(* Logix 5000 project; controller PLC_MCC1201_220AP1 vendor 1 type 14 code 164 rev 35.11; software revision 35.00; part 13 of 25 *)
(* tags used below, declared in another part *)
   B180 : DINT[10];
   B3 : DINT[102];
   BIN_1B_EAST : ALIAS FOR O[112].12;
   BT181_000 : MESSAGE;
   BT181_001 : MESSAGE;
   BT181_002 : MESSAGE;
   BT181_003 : MESSAGE;
   C1_PNL_FLT : ALIAS FOR I[113].2;
   C2_PNL_FLT : ALIAS FOR I[113].3;
   C3_PNL_FLT : ALIAS FOR I[113].4;
   C4_PNL_FLT : ALIAS FOR I[113].1;
   C5 : COUNTER[100];
   CAP_ALM_HORN : ALIAS FOR O[11].2;
   CR1_DOWN_PROX : ALIAS FOR I[64].11;
   CR1_RUN_ENABLE : ALIAS FOR O[117].4;
   CULL_FLT : ALIAS FOR B3[3].1;
   CULLET_FLT_PL : ALIAS FOR O[11].1;
   DIV_POSITION : ALIAS FOR I[24].12;
   I : INT[128];
   LEG2_SLEEP : ALIAS FOR I[123].14;
   LEG3_SLEEP : ALIAS FOR I[123].15;
   LEG4_SLEEP : ALIAS FOR I[124].0;
   LEG5_SLEEP : ALIAS FOR I[124].1;
   M37B_FWD_DIR : ALIAS FOR B3[1].14;
   M37B_FWD_PL : ALIAS FOR O[25].5;
   M37B_FWD_SIG : ALIAS FOR I[112].3;
   M37B_FWD_SS : ALIAS FOR I[24].8;
   M37B_REV_DIR : ALIAS FOR B3[1].15;
   M37B_REV_PL : ALIAS FOR O[25].6;
   M37B_REV_SIG : ALIAS FOR I[112].4;
   M37B_REV_SS : ALIAS FOR I[24].9;
   M37B_RUN_FWD : ALIAS FOR O[119].0;
   M37B_RUN_REV : ALIAS FOR O[119].1;
   M47_REV_SS : ALIAS FOR I[24].11;
   M47B_FWD_DIR : ALIAS FOR B3[1].12;
   M47B_FWD_PL : ALIAS FOR O[25].7;
   M47B_FWD_SIG : ALIAS FOR I[112].1;
   M47B_FWD_SS : ALIAS FOR I[24].10;
   M47B_REV_DIR : ALIAS FOR B3[1].13;
   M47B_REV_PL : ALIAS FOR O[25].8;
   M47B_REV_SIG : ALIAS FOR I[112].2;
   M47B_RUN_FWD : ALIAS FOR O[119].2;
   M47B_RUN_REV : ALIAS FOR O[119].3;
   N53 : DINT[10];
   N54 : DINT[501];
   N60 : DINT[420];
   O : INT[128];
   REL_DRV_FLT : ALIAS FOR B3[3].0;
   RELIANCE_FLT_PL : ALIAS FOR O[11].0;
   S : INT[128];
   SPNGE_DN_FLT : ALIAS FOR I[43].5;
   SPNGE_UP_FLT : ALIAS FOR I[43].4;
   Status : INT;   // INT tag to retrieve Status value through GSV created during conversion
   T4 : TIMER[100];
   T51 : TIMER[13];
   TMP_xAlwaysOFF : BOOL;
   TONY : ALIAS FOR B3[10].15;
   VMCCMB_ALM_HRN : ALIAS FOR O[20].3;
   VP917060_MED : ALIAS FOR O[116].14;
   VP917060_THICK : ALIAS FOR O[116].15;
   VP917060_THIN : ALIAS FOR O[116].13;
   VP917065_MED : ALIAS FOR O[114].5;
   VP917065_THICK : ALIAS FOR O[114].6;
   VP917065_THIN : ALIAS FOR O[114].4;
   VP917066_MED : ALIAS FOR O[114].2;
   VP917066_THICK : ALIAS FOR O[114].3;
   VP917066_THIN : ALIAS FOR O[114].1;
   VP917067_MED : ALIAS FOR O[113].15;
   VP917067_THICK : ALIAS FOR O[114].0;
   VP917067_THIN : ALIAS FOR O[113].14;
   VP917070_MED : ALIAS FOR O[114].8;
   VP917070_THICK : ALIAS FOR O[114].9;
   VP917070_THIN : ALIAS FOR O[114].7;
   VP917071_MED : ALIAS FOR O[114].11;
   VP917071_THICK : ALIAS FOR O[114].12;
   VP917071_THIN : ALIAS FOR O[114].10;
   VP917072_MED : ALIAS FOR O[116].11;
   VP917072_THICK : ALIAS FOR O[116].12;
   VP917072_THIN : ALIAS FOR O[116].10;
   VP917073_MED : ALIAS FOR O[115].14;
   VP917073_THICK : ALIAS FOR O[115].15;
   VP917073_THIN : ALIAS FOR O[115].13;
   VP917074_MED : ALIAS FOR O[115].11;
   VP917074_THICK : ALIAS FOR O[115].12;
   VP917074_THIN : ALIAS FOR O[115].10;
   VP917075_MED : ALIAS FOR O[115].8;
   VP917075_THICK : ALIAS FOR O[115].9;
   VP917075_THIN : ALIAS FOR O[115].7;
   VP917076_MED : ALIAS FOR O[115].5;
   VP917076_THICK : ALIAS FOR O[115].6;
   VP917076_THIN : ALIAS FOR O[115].4;
   VP917077_MED : ALIAS FOR O[114].14;
   VP917077_THICK : ALIAS FOR O[114].15;
   VP917077_THIN : ALIAS FOR O[114].13;
   W1_DRV_FLT_RES : ALIAS FOR O[47].2;
(* MainProgram, continued *)

ROUTINE _107_LADDER   (* ladder *)
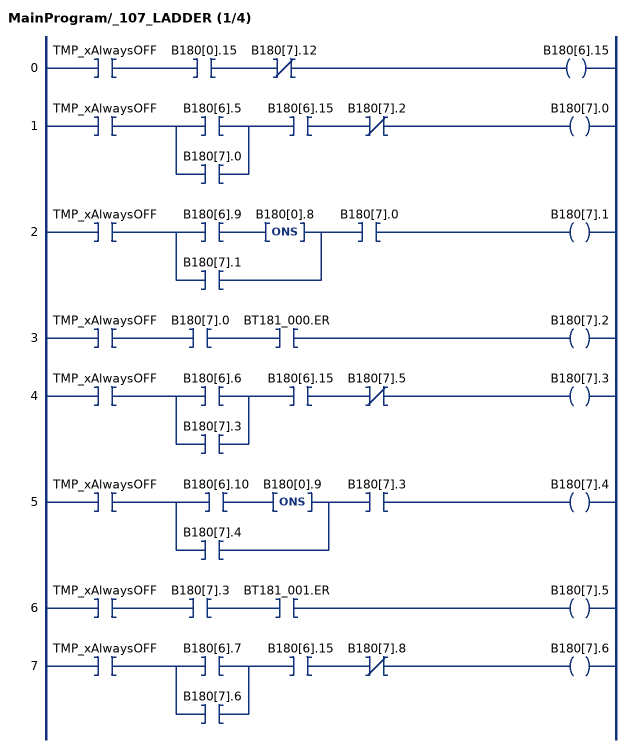
   0: XIC(TMP_xAlwaysOFF)XIC(B180[0].15)XIO(B180[7].12)OTE(B180[6].15);
   1: XIC(TMP_xAlwaysOFF)[XIC(B180[6].5) ,XIC(B180[7].0) ]XIC(B180[6].15)XIO(B180[7].2)OTE(B180[7].0);
   2: XIC(TMP_xAlwaysOFF)[XIC(B180[6].9) ONS(B180[0].8) ,XIC(B180[7].1) ]XIC(B180[7].0)OTE(B180[7].1);
   3: XIC(TMP_xAlwaysOFF)XIC(B180[7].0)XIC(BT181_000.ER)OTE(B180[7].2);
   4: XIC(TMP_xAlwaysOFF)[XIC(B180[6].6) ,XIC(B180[7].3) ]XIC(B180[6].15)XIO(B180[7].5)OTE(B180[7].3);
   5: XIC(TMP_xAlwaysOFF)[XIC(B180[6].10) ONS(B180[0].9) ,XIC(B180[7].4) ]XIC(B180[7].3)OTE(B180[7].4);
   6: XIC(TMP_xAlwaysOFF)XIC(B180[7].3)XIC(BT181_001.ER)OTE(B180[7].5);
   7: XIC(TMP_xAlwaysOFF)[XIC(B180[6].7) ,XIC(B180[7].6) ]XIC(B180[6].15)XIO(B180[7].8)OTE(B180[7].6);
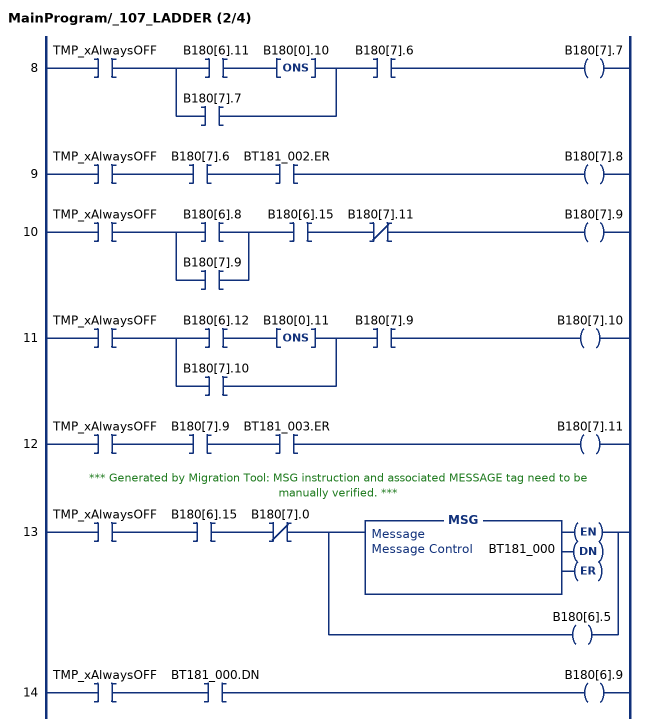
   8: XIC(TMP_xAlwaysOFF)[XIC(B180[6].11) ONS(B180[0].10) ,XIC(B180[7].7) ]XIC(B180[7].6)OTE(B180[7].7);
   9: XIC(TMP_xAlwaysOFF)XIC(B180[7].6)XIC(BT181_002.ER)OTE(B180[7].8);
   10: XIC(TMP_xAlwaysOFF)[XIC(B180[6].8) ,XIC(B180[7].9) ]XIC(B180[6].15)XIO(B180[7].11)OTE(B180[7].9);
   11: XIC(TMP_xAlwaysOFF)[XIC(B180[6].12) ONS(B180[0].11) ,XIC(B180[7].10) ]XIC(B180[7].9)OTE(B180[7].10);
   12: XIC(TMP_xAlwaysOFF)XIC(B180[7].9)XIC(BT181_003.ER)OTE(B180[7].11);
   // *** Generated by Migration Tool: MSG instruction and associated MESSAGE tag need to be manually verified. ***
   13: XIC(TMP_xAlwaysOFF)XIC(B180[6].15)XIO(B180[7].0)[MSG(BT181_000) ,OTE(B180[6].5) ];
   14: XIC(TMP_xAlwaysOFF)XIC(BT181_000.DN)OTE(B180[6].9);
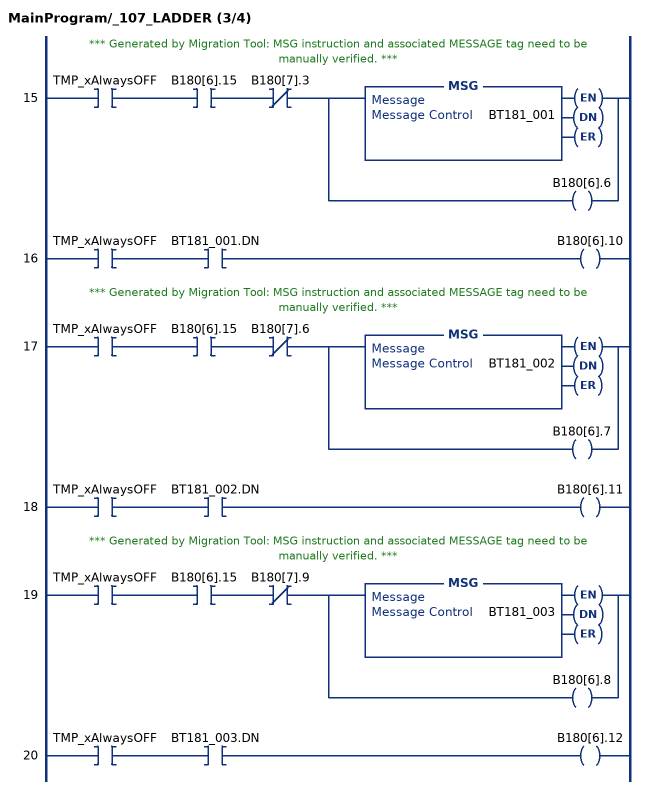
   // *** Generated by Migration Tool: MSG instruction and associated MESSAGE tag need to be manually verified. ***
   15: XIC(TMP_xAlwaysOFF)XIC(B180[6].15)XIO(B180[7].3)[MSG(BT181_001) ,OTE(B180[6].6) ];
   16: XIC(TMP_xAlwaysOFF)XIC(BT181_001.DN)OTE(B180[6].10);
   // *** Generated by Migration Tool: MSG instruction and associated MESSAGE tag need to be manually verified. ***
   17: XIC(TMP_xAlwaysOFF)XIC(B180[6].15)XIO(B180[7].6)[MSG(BT181_002) ,OTE(B180[6].7) ];
   18: XIC(TMP_xAlwaysOFF)XIC(BT181_002.DN)OTE(B180[6].11);
   // *** Generated by Migration Tool: MSG instruction and associated MESSAGE tag need to be manually verified. ***
   19: XIC(TMP_xAlwaysOFF)XIC(B180[6].15)XIO(B180[7].9)[MSG(BT181_003) ,OTE(B180[6].8) ];
   20: XIC(TMP_xAlwaysOFF)XIC(BT181_003.DN)OTE(B180[6].12);
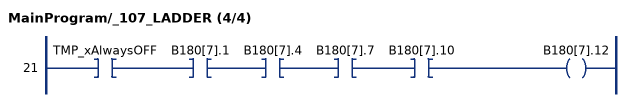
   21: XIC(TMP_xAlwaysOFF)XIC(B180[7].1)XIC(B180[7].4)XIC(B180[7].7)XIC(B180[7].10)OTE(B180[7].12);
END_ROUTINE

ROUTINE _10_SLEEP   (* ladder *)
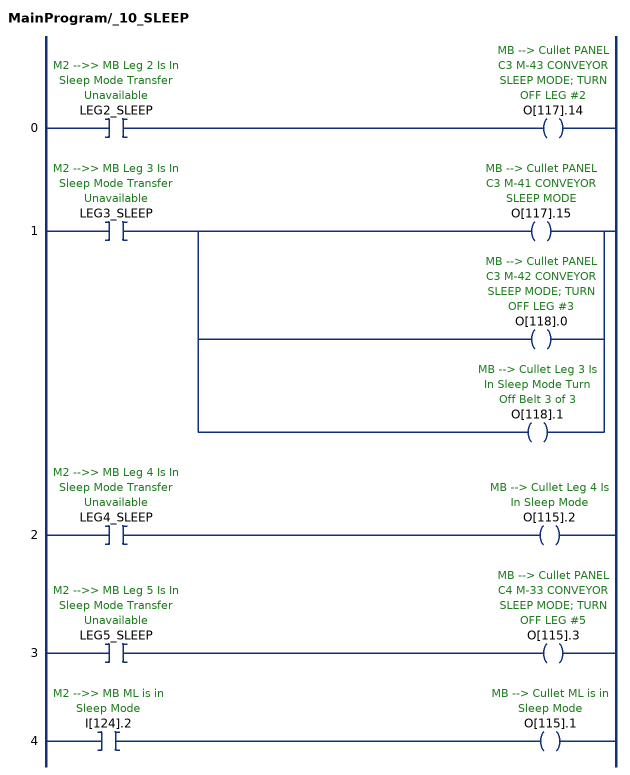
   0: XIC(LEG2_SLEEP)OTE(O[117].14);
   1: XIC(LEG3_SLEEP)[OTE(O[117].15) ,OTE(O[118].0) ,OTE(O[118].1) ];
   2: XIC(LEG4_SLEEP)OTE(O[115].2);
   3: XIC(LEG5_SLEEP)OTE(O[115].3);
   4: XIC(I[124].2)OTE(O[115].1);
END_ROUTINE

ROUTINE _11_CULLET   (* ladder *)
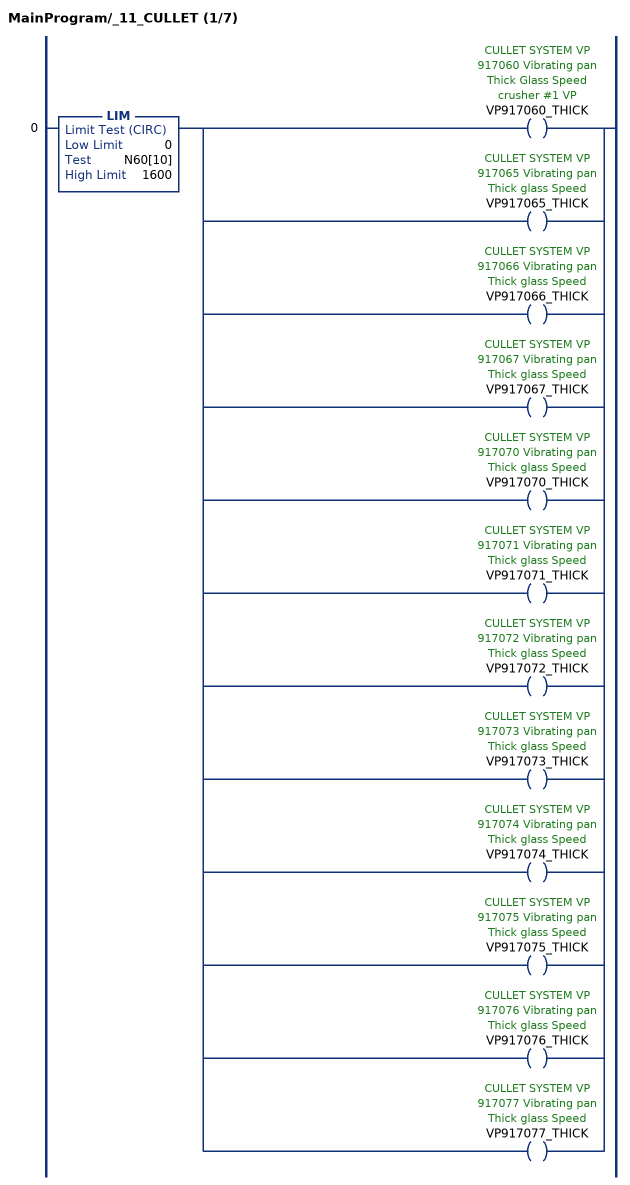
   0: LIM(0,N60[10],1600)[OTE(VP917060_THICK) ,OTE(VP917065_THICK) ,OTE(VP917066_THICK) ,OTE(VP917067_THICK) ,OTE(VP917070_THICK) ,OTE(VP917071_THICK) ,OTE(VP917072_THICK) ,OTE(VP917073_THICK) ,OTE(VP917074_THICK) ,OTE(VP917075_THICK) ,OTE(VP917076_THICK) ,OTE(VP917077_THICK) ];
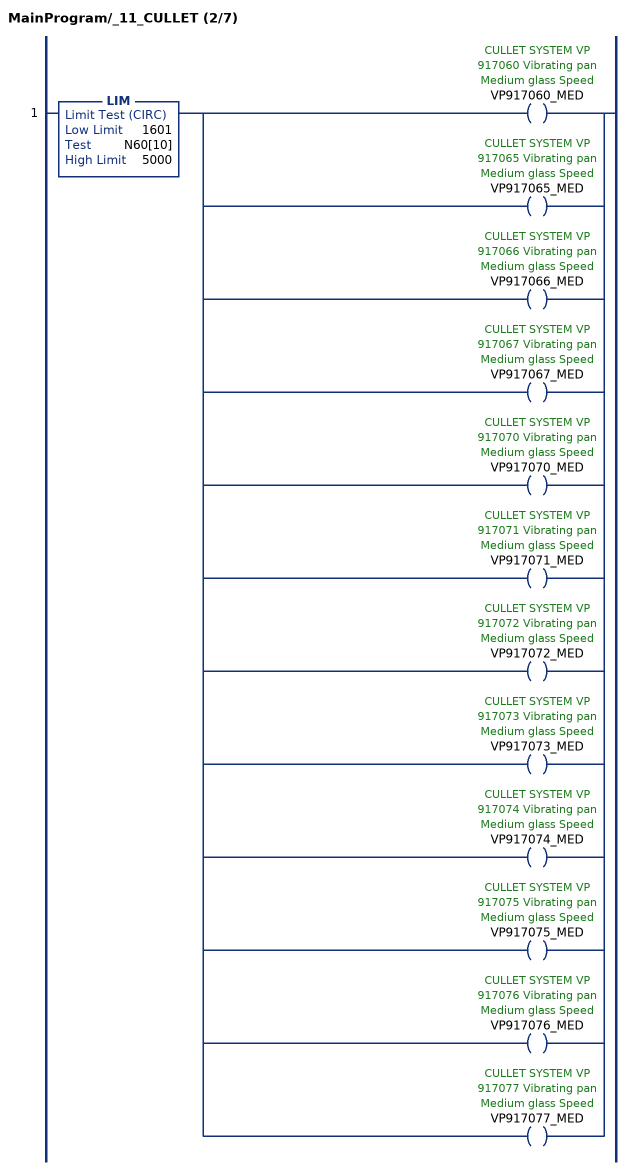
   1: LIM(1601,N60[10],5000)[OTE(VP917060_MED) ,OTE(VP917065_MED) ,OTE(VP917066_MED) ,OTE(VP917067_MED) ,OTE(VP917070_MED) ,OTE(VP917071_MED) ,OTE(VP917072_MED) ,OTE(VP917073_MED) ,OTE(VP917074_MED) ,OTE(VP917075_MED) ,OTE(VP917076_MED) ,OTE(VP917077_MED) ];
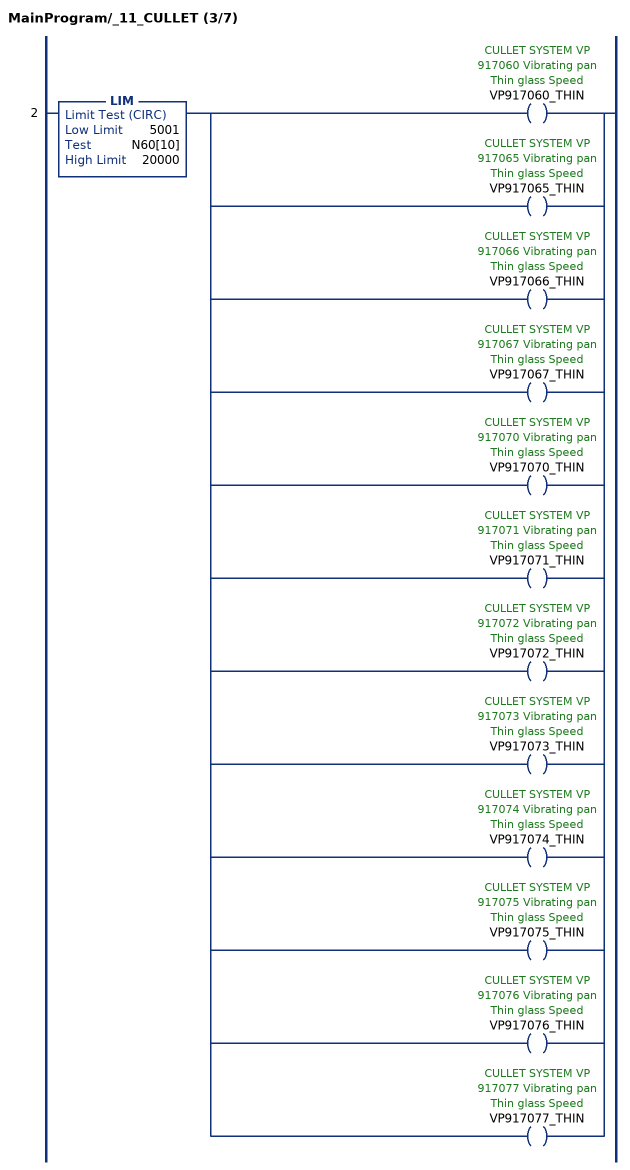
   2: LIM(5001,N60[10],20000)[OTE(VP917060_THIN) ,OTE(VP917065_THIN) ,OTE(VP917066_THIN) ,OTE(VP917067_THIN) ,OTE(VP917070_THIN) ,OTE(VP917071_THIN) ,OTE(VP917072_THIN) ,OTE(VP917073_THIN) ,OTE(VP917074_THIN) ,OTE(VP917075_THIN) ,OTE(VP917076_THIN) ,OTE(VP917077_THIN) ];
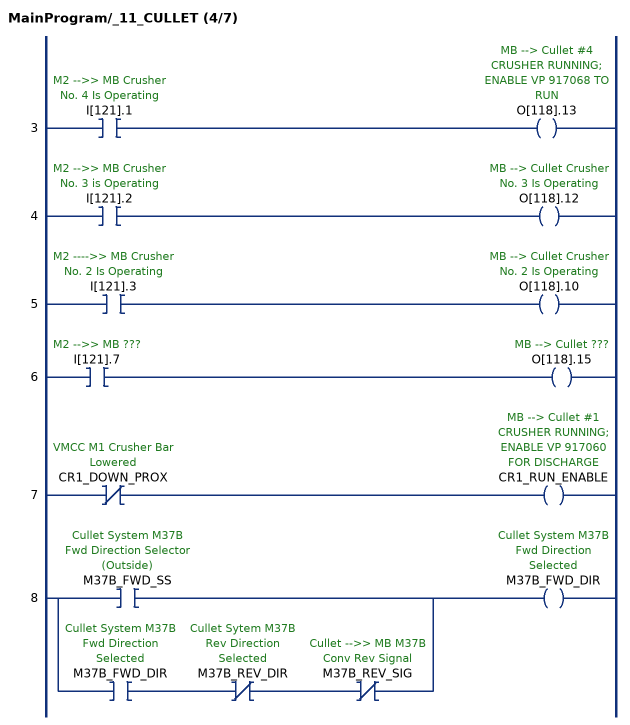
   3: XIC(I[121].1)OTE(O[118].13);
   4: XIC(I[121].2)OTE(O[118].12);
   5: XIC(I[121].3)OTE(O[118].10);
   6: XIC(I[121].7)OTE(O[118].15);
   7: XIO(CR1_DOWN_PROX)OTE(CR1_RUN_ENABLE);
   8: [XIC(M37B_FWD_SS) ,XIC(M37B_FWD_DIR) XIO(M37B_REV_DIR) XIO(M37B_REV_SIG) ]OTE(M37B_FWD_DIR);
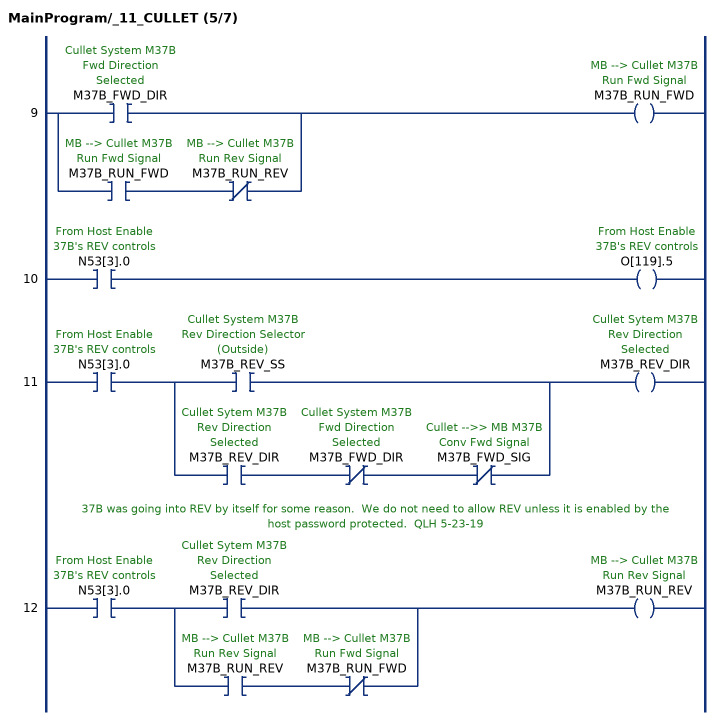
   9: [XIC(M37B_FWD_DIR) ,XIC(M37B_RUN_FWD) XIO(M37B_RUN_REV) ]OTE(M37B_RUN_FWD);
   10: XIC(N53[3].0)OTE(O[119].5);
   11: XIC(N53[3].0)[XIC(M37B_REV_SS) ,XIC(M37B_REV_DIR) XIO(M37B_FWD_DIR) XIO(M37B_FWD_SIG) ]OTE(M37B_REV_DIR);
   // 37B was going into REV by itself for some reason.  We do not need to allow REV unless it is enabled by the host password protected.  QLH 5-23-19
   12: XIC(N53[3].0)[XIC(M37B_REV_DIR) ,XIC(M37B_RUN_REV) XIO(M37B_RUN_FWD) ]OTE(M37B_RUN_REV);
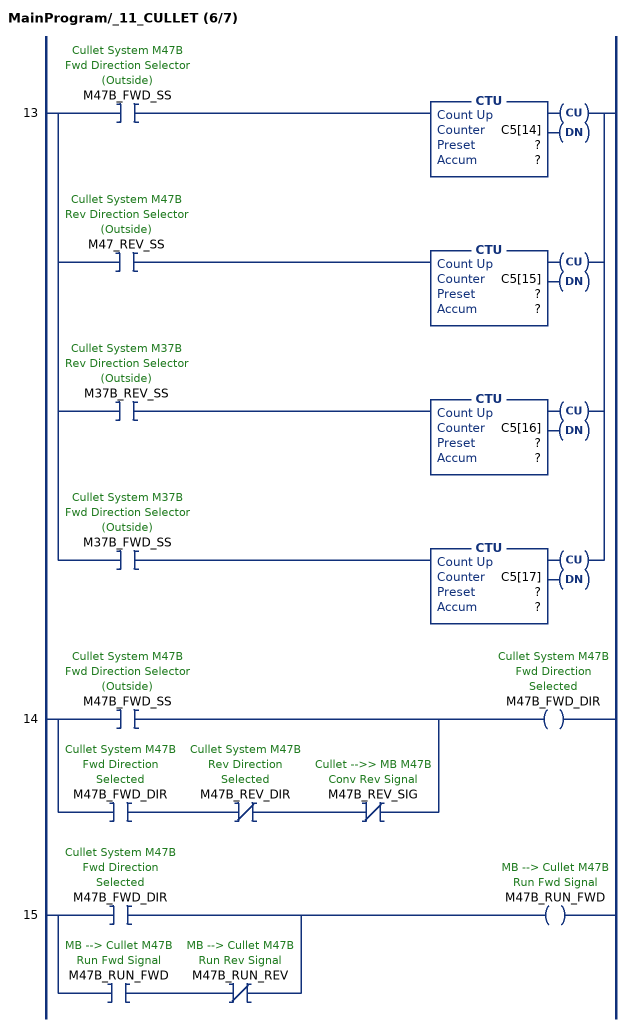
   13: [XIC(M47B_FWD_SS) CTU(C5[14],?,?) ,XIC(M47_REV_SS) CTU(C5[15],?,?) ,XIC(M37B_REV_SS) CTU(C5[16],?,?) ,XIC(M37B_FWD_SS) CTU(C5[17],?,?) ];
   14: [XIC(M47B_FWD_SS) ,XIC(M47B_FWD_DIR) XIO(M47B_REV_DIR) XIO(M47B_REV_SIG) ]OTE(M47B_FWD_DIR);
   15: [XIC(M47B_FWD_DIR) ,XIC(M47B_RUN_FWD) XIO(M47B_RUN_REV) ]OTE(M47B_RUN_FWD);
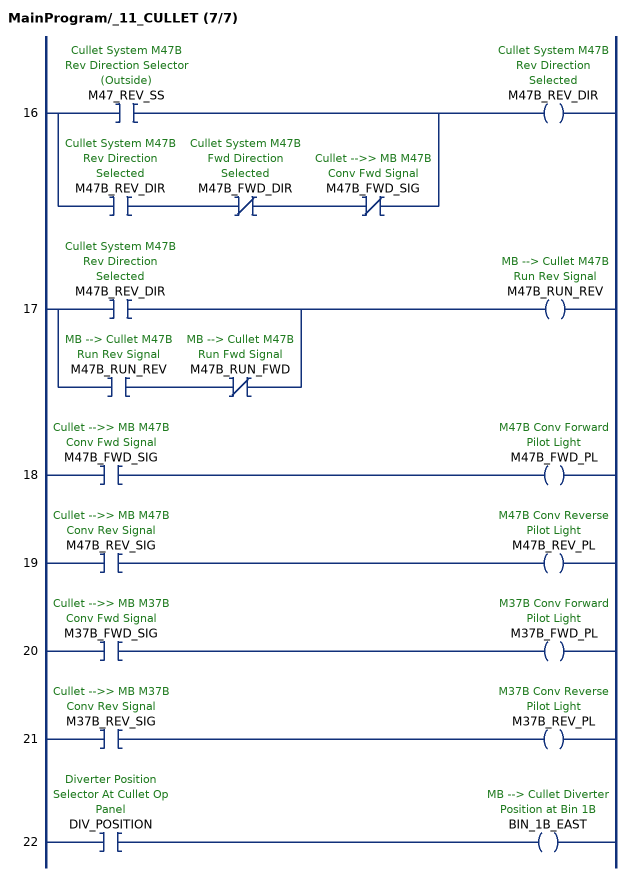
   16: [XIC(M47_REV_SS) ,XIC(M47B_REV_DIR) XIO(M47B_FWD_DIR) XIO(M47B_FWD_SIG) ]OTE(M47B_REV_DIR);
   17: [XIC(M47B_REV_DIR) ,XIC(M47B_RUN_REV) XIO(M47B_RUN_FWD) ]OTE(M47B_RUN_REV);
   18: XIC(M47B_FWD_SIG)OTE(M47B_FWD_PL);
   19: XIC(M47B_REV_SIG)OTE(M47B_REV_PL);
   20: XIC(M37B_FWD_SIG)OTE(M37B_FWD_PL);
   21: XIC(M37B_REV_SIG)OTE(M37B_REV_PL);
   22: XIC(DIV_POSITION)OTE(BIN_1B_EAST);
END_ROUTINE

ROUTINE _12_MAIN   (* ladder *)
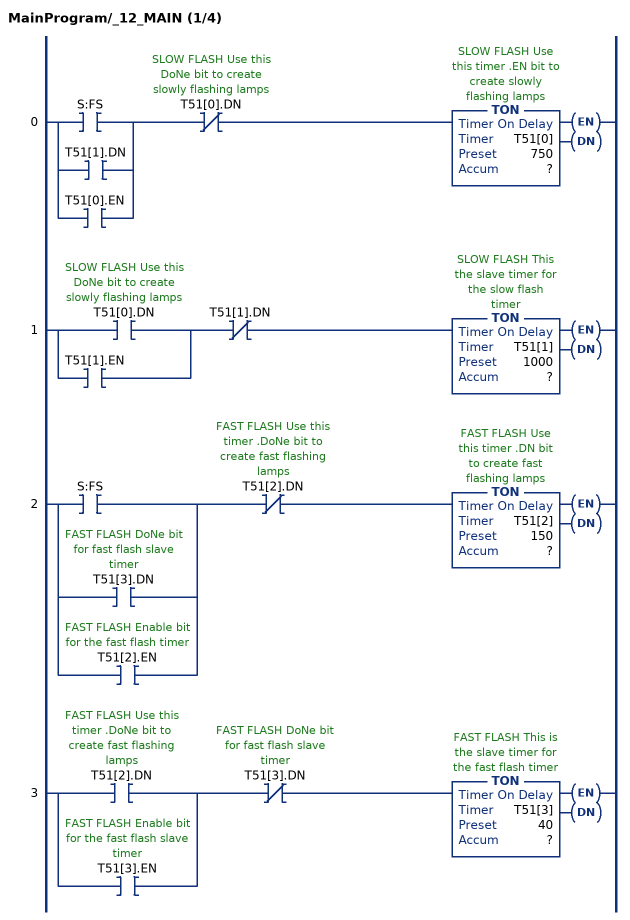
   0: [XIC(S:FS) ,XIC(T51[1].DN) ,XIC(T51[0].EN) ]XIO(T51[0].DN)TON(T51[0],?,?);
   1: [XIC(T51[0].DN) ,XIC(T51[1].EN) ]XIO(T51[1].DN)TON(T51[1],?,?);
   2: [XIC(S:FS) ,XIC(T51[3].DN) ,XIC(T51[2].EN) ]XIO(T51[2].DN)TON(T51[2],?,?);
   3: [XIC(T51[2].DN) ,XIC(T51[3].EN) ]XIO(T51[3].DN)TON(T51[3],?,?);
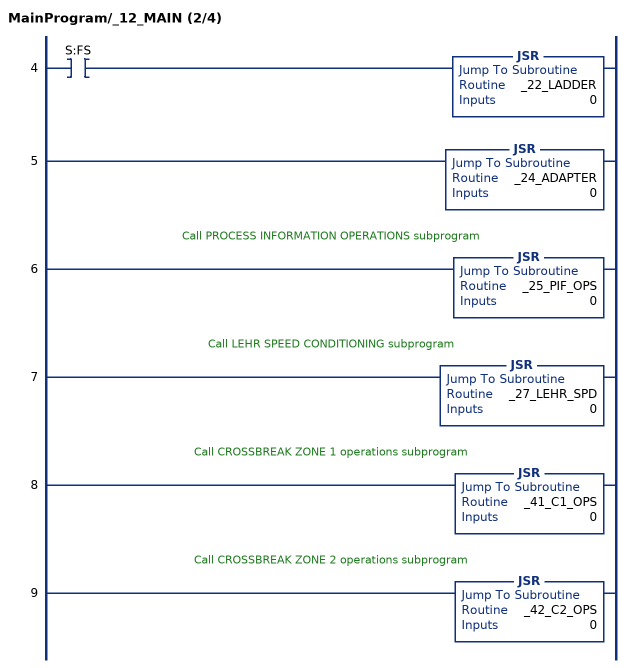
   4: XIC(S:FS)JSR(_22_LADDER,0);
   5: JSR(_24_ADAPTER,0);
   // Call PROCESS INFORMATION OPERATIONS subprogram
   6: JSR(_25_PIF_OPS,0);
   // Call LEHR SPEED CONDITIONING subprogram
   7: JSR(_27_LEHR_SPD,0);
   // Call CROSSBREAK ZONE 1 operations subprogram
   8: JSR(_41_C1_OPS,0);
   // Call CROSSBREAK ZONE 2 operations subprogram
   9: JSR(_42_C2_OPS,0);
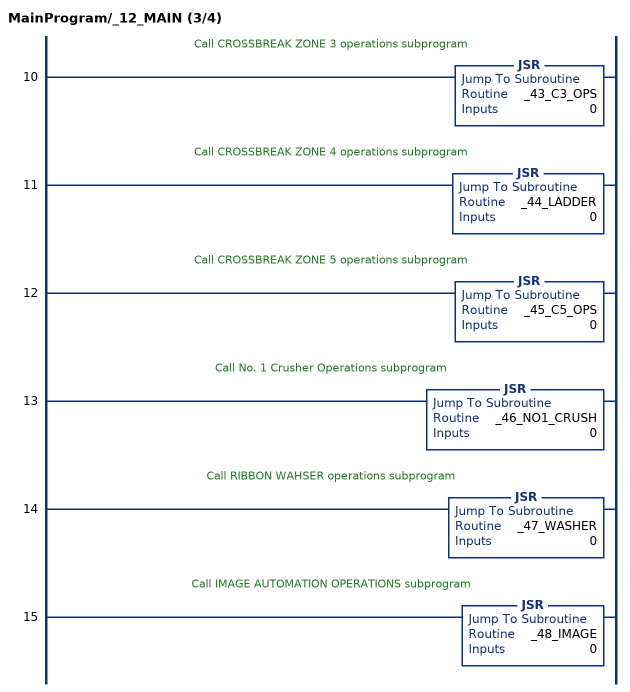
   // Call CROSSBREAK ZONE 3 operations subprogram
   10: JSR(_43_C3_OPS,0);
   // Call CROSSBREAK ZONE 4 operations subprogram
   11: JSR(_44_LADDER,0);
   // Call CROSSBREAK ZONE 5 operations subprogram
   12: JSR(_45_C5_OPS,0);
   // Call No. 1 Crusher Operations subprogram
   13: JSR(_46_NO1_CRUSH,0);
   // Call RIBBON WAHSER operations subprogram
   14: JSR(_47_WASHER,0);
   // Call IMAGE AUTOMATION OPERATIONS subprogram
   15: JSR(_48_IMAGE,0);
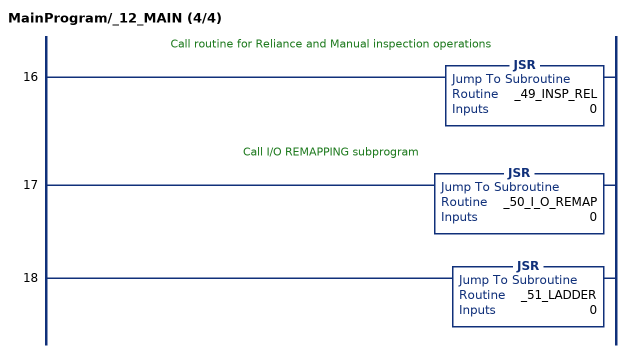
   // Call routine for Reliance and Manual inspection operations
   16: JSR(_49_INSP_REL,0);
   // Call I/O REMAPPING subprogram
   17: JSR(_50_I_O_REMAP,0);
   18: JSR(_51_LADDER,0);
END_ROUTINE

ROUTINE _13_ALARMING   (* ladder *)
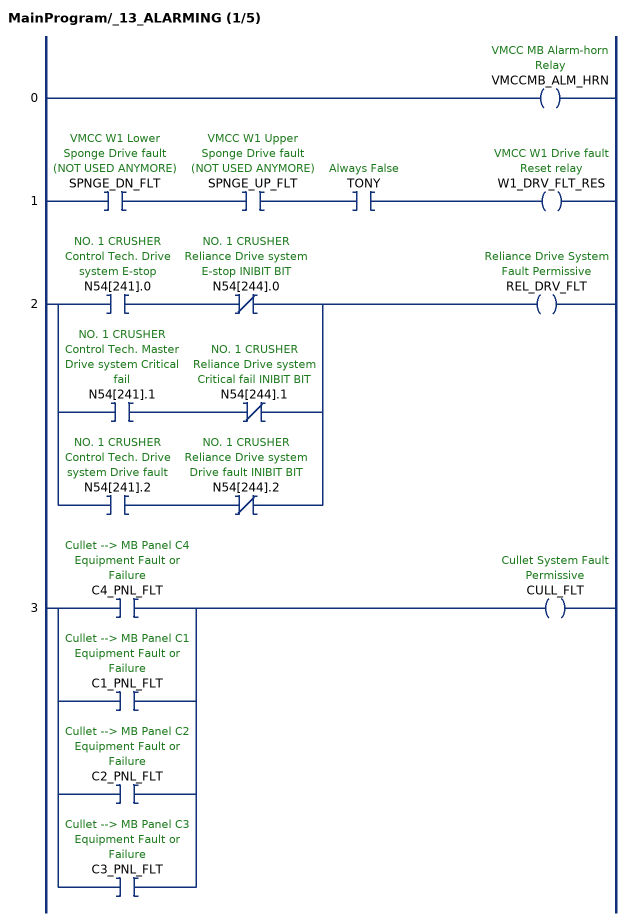
   0: OTE(VMCCMB_ALM_HRN);
   1: XIC(SPNGE_DN_FLT)XIC(SPNGE_UP_FLT)XIC(TONY)OTE(W1_DRV_FLT_RES);
   2: [XIC(N54[241].0) XIO(N54[244].0) ,XIC(N54[241].1) XIO(N54[244].1) ,XIC(N54[241].2) XIO(N54[244].2) ]OTE(REL_DRV_FLT);
   3: [XIC(C4_PNL_FLT) ,XIC(C1_PNL_FLT) ,XIC(C2_PNL_FLT) ,XIC(C3_PNL_FLT) ]OTE(CULL_FLT);
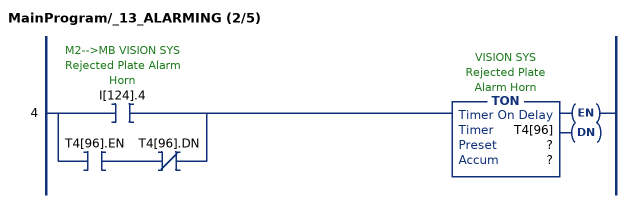
   4: [XIC(I[124].4) ,XIC(T4[96].EN) XIO(T4[96].DN) ]TON(T4[96],?,?);
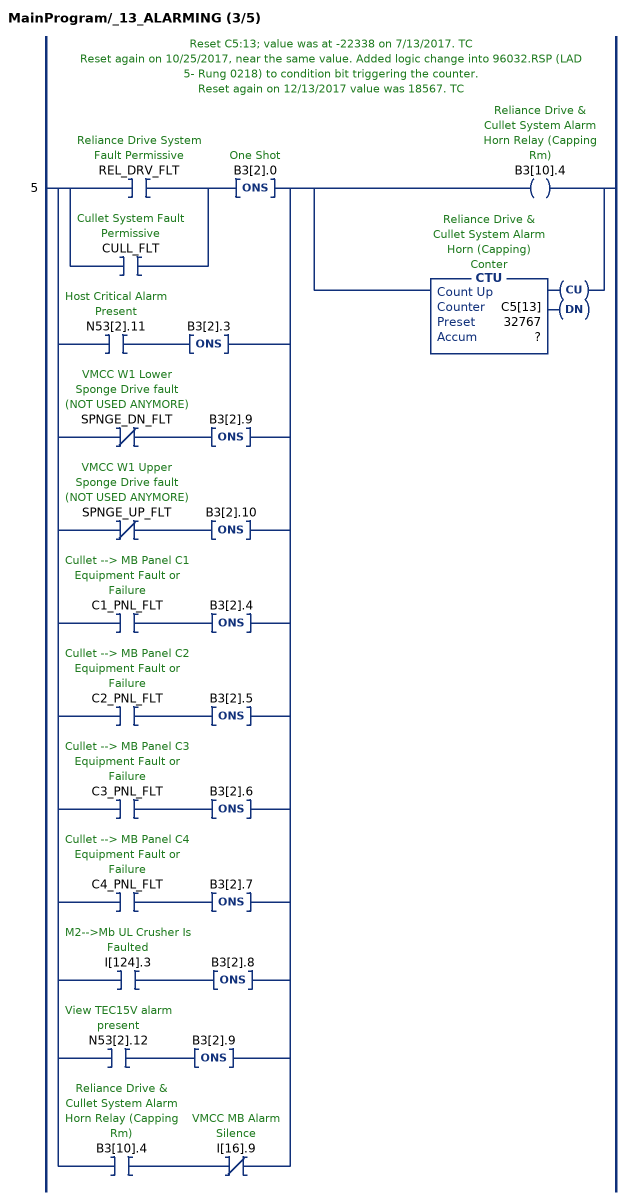
   // Reset C5:13; value was at -22338 on 7/13/2017. TC
   //                                                                                                                                                                     Reset again on 10/25/2017, near the same value. Added logic change into 96032.RSP (LAD 5- Rung 0218) to condition bit triggering the counter.
   //                                                                                                                                                                                                                  Reset again on 12/13/2017 value was 18567. TC
   5: [[[XIC(REL_DRV_FLT) ,XIC(CULL_FLT) ] ONS(B3[2].0) ,XIC(N53[2].11) ONS(B3[2].3) ,XIO(SPNGE_DN_FLT) ONS(B3[2].9) ,XIO(SPNGE_UP_FLT) ONS(B3[2].10) ,XIC(C1_PNL_FLT) ONS(B3[2].4) ,XIC(C2_PNL_FLT) ONS(B3[2].5) ,XIC(C3_PNL_FLT) ONS(B3[2].6) ,XIC(C4_PNL_FLT) ONS(B3[2].7) ,XIC(I[124].3) ONS(B3[2].8) ,XIC(N53[2].12) ONS(B3[2].9) ] ,XIC(B3[10].4) XIO(I[16].9) ][OTE(B3[10].4) ,CTU(C5[13],?,?) ];
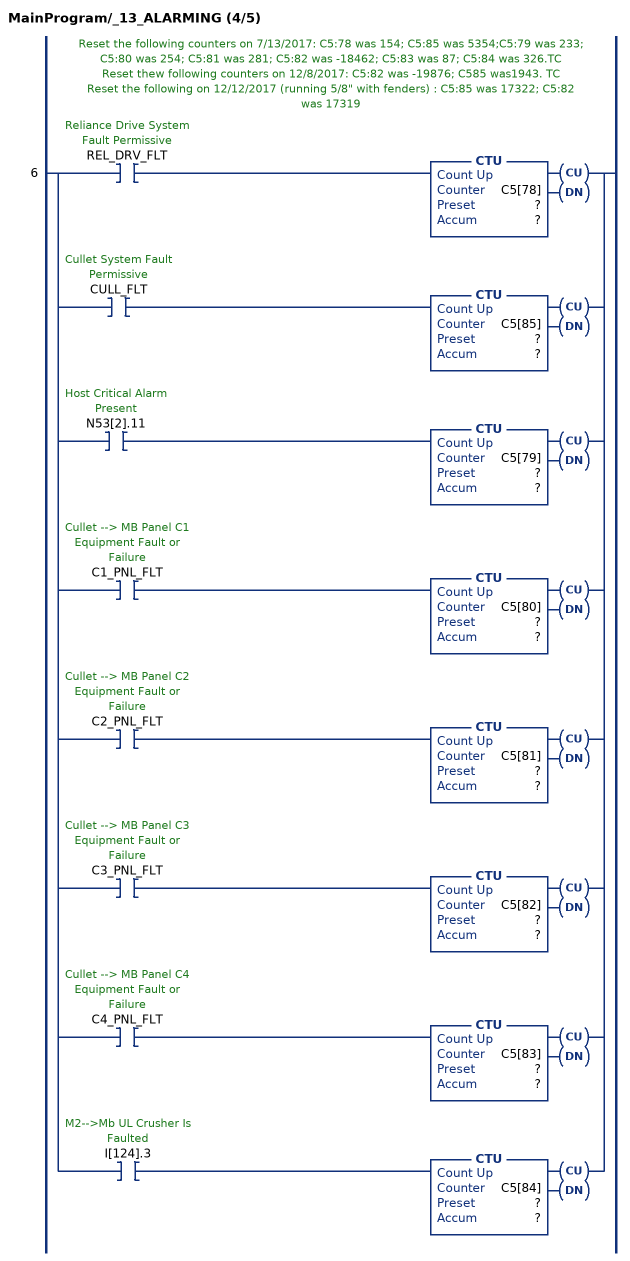
   // Reset the following counters on 7/13/2017: C5:78 was 154; C5:85 was 5354;C5:79 was 233; C5:80 was 254; C5:81 was 281; C5:82 was -18462; C5:83 was 87; C5:84 was 326.TC
   //                                                                                                                       Reset thew following counters on 12/8/2017: C5:82 was -19876; C585 was1943. TC
   //                                                                                                                       Reset the following on 12/12/2017 (running 5/8" with fenders) : C5:85 was 17322; C5:82 was 17319
   6: [[XIC(REL_DRV_FLT) CTU(C5[78],?,?) ,XIC(CULL_FLT) CTU(C5[85],?,?) ] ,XIC(N53[2].11) CTU(C5[79],?,?) ,XIC(C1_PNL_FLT) CTU(C5[80],?,?) ,XIC(C2_PNL_FLT) CTU(C5[81],?,?) ,XIC(C3_PNL_FLT) CTU(C5[82],?,?) ,XIC(C4_PNL_FLT) CTU(C5[83],?,?) ,XIC(I[124].3) CTU(C5[84],?,?) ];
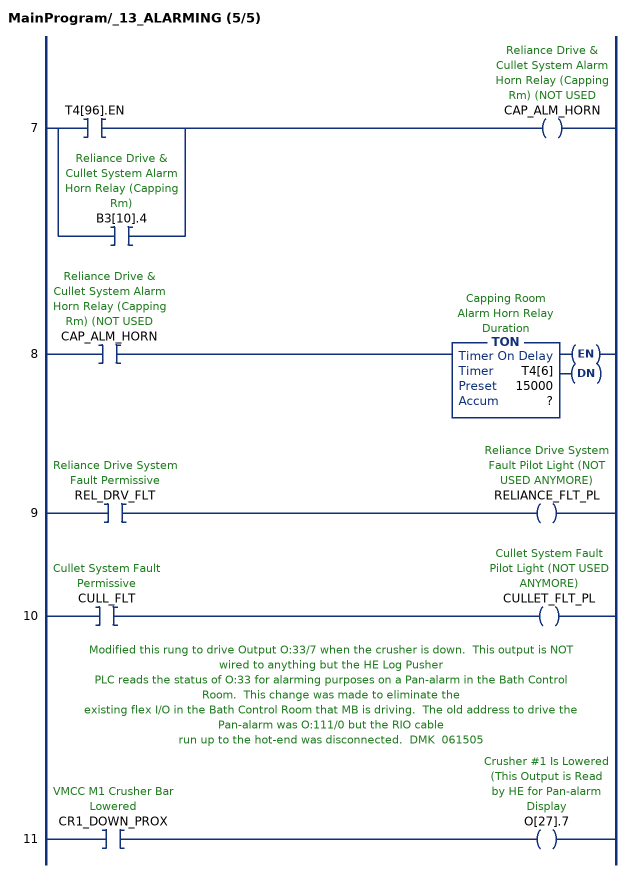
   7: [XIC(T4[96].EN) ,XIC(B3[10].4) ]OTE(CAP_ALM_HORN);
   8: XIC(CAP_ALM_HORN)TON(T4[6],?,?);
   9: XIC(REL_DRV_FLT)OTE(RELIANCE_FLT_PL);
   10: XIC(CULL_FLT)OTE(CULLET_FLT_PL);
   // Modified this rung to drive Output O:33/7 when the crusher is down.  This output is NOT wired to anything but the HE Log Pusher
   // PLC reads the status of O:33 for alarming purposes on a Pan-alarm in the Bath Control Room.  This change was made to eliminate the
   // existing flex I/O in the Bath Control Room that MB is driving.  The old address to drive the Pan-alarm was O:111/0 but the RIO cable
   // run up to the hot-end was disconnected.  DMK  061505
   11: XIC(CR1_DOWN_PROX)OTE(O[27].7);
END_ROUTINE
